
           "RPA30_DataBlock".RPA30_show_points_hmi := 0;
           "RPA30_DataBlock".RPA30_UseInterval_Primer207 := false;
           "RPA30_DataBlock".RPA30_UseIntervalBottleRemover208 := false;
           "RPA30_DataBlock".RPA30_cyclusState := "RPA30_go_to_home_position";
       END_IF;

       "RPA30_DataBlock".RPA30_actual_instruction_index := 255;

       "RPA30R_Beacon_1_LCDPanelGreen" := false;
       "RPA30R_Beacon_1_LCDPanelOrange" := false;
       "RPA30R_Beacon_1_LCDPanelRed" := false;
       "RPA30R_Beacon_1_LCDPanelSiren" := false;
       "RPA30R_Beacon_2_PrimerBoxGreen" := false;
       "RPA30R_Beacon_2_PrimerBoxOrange" := false;
       "RPA30R_Beacon_2_PrimerBoxRed" := false;
       "RPA30R_Beacon_2_PrimerBoxSiren" := false;

       "RPA30R_PrimerPA30GreenReady" := false;
       "RPA30R_PrimerPA30GreenFelt" := false;
       "RPA30R_PrimerPA30GreenRemover208" := false;
       "RPA30R_PrimerPA30GreenPrimer207" := false;
       "RPA30R_PrimerPA30RedNotReady" := false;
       "RPA30R_PrimerPA30RedChangePad" := false;
       "RPA30R_LedBlueConfirm" := false;
       "RPA30R_light" := false;

       "RPA30_DataBlock".RPA30_scannedFrameBareCode := '';

       //if station not active
       "StartStation"(startButton := "RPA30R_LCDButtonStart",
                      StationStartControlVariable := "RPA30_DataBlock".RPA30_Start,
                      stationLight := "RPA30R_light");

       "startButtonLightControlHandler"(stationActivitycontrolVariable := "RPA30_DataBlock".RPA30_Start,
                                        startButtonLED := "RPA30R_LEDGreenSart");
   END_IF;



   IF "RPA30_DataBlock".RPA30_state_information_send = true THEN
       "RPA30_DataBlock".RPA30_state_information_send := NOT "pa30r_station_monitoring"(station_configuration := "RPA30_DataBlock".RPA30_station_configuration,
                                                                                       fail_state := "RPA30_DataBlock".RPA30_failStateLock,
                                                                                       big_fail_state := "RPA30_DataBlock".RPA30_bigFailStateLock,
                                                                                       error_state := "RPA30_DataBlock".RPA30_ErrorStateLock,
                                                                                       fatal_error_state := "RPA30_DataBlock".RPA30_fatalErrorStateLock,
                                                                                       work_cyclus_state := "RPA30_DataBlock".RPA30_actual_instruction_index,
                                                                                       current_frame_code := "RPA30_DataBlock".RPA30_scannedFrameBareCode,
                                                                                       station_activity_state := "RPA30_DataBlock".RPA30_Start,
                                                                                       position_sensor_y := "RPA30R_RoofRotationSensorYAtOperator",
                                                                                       server_connection := "tcp_datablock".tcp_connection,
                                                                                       index:="tcp_datablock".pa30r_station_state_index);
   ELSE
       IF "RPA30_DataBlock".RPA30_fail_state_pre <> "RPA30_DataBlock".RPA30_failStateLock OR
           "RPA30_DataBlock".RPA30_error_state_pre <> "RPA30_DataBlock".RPA30_ErrorStateLock OR
           "RPA30_DataBlock".RPA30_big_fail_state_pre <> "RPA30_DataBlock".RPA30_bigFailStateLock OR
           "RPA30_DataBlock".RPA30_fatal_error_state_pre <> "RPA30_DataBlock".RPA30_fatalErrorStateLock OR
           "RPA30_DataBlock".RPA30_current_frame_code_pre <> "RPA30_DataBlock".RPA30_scannedFrameBareCode OR
           "RPA30_DataBlock".RPA30_hmi_state_pre <> "RPA30_DataBlock".RPA30_actual_instruction_index OR
           "RPA30_DataBlock".RPA30_position_y_pre <> "RPA30R_RoofRotationSensorYAtOperator" OR
           "RPA30_DataBlock".RPA30_station_activity_state_pre <> "RPA30_DataBlock".RPA30_Start THEN

           "RPA30_DataBlock".RPA30_state_information_send := true;
       END_IF;

       "RPA30_DataBlock".RPA30_fail_state_pre := "RPA30_DataBlock".RPA30_failStateLock;
       "RPA30_DataBlock".RPA30_error_state_pre := "RPA30_DataBlock".RPA30_ErrorStateLock;
       "RPA30_DataBlock".RPA30_big_fail_state_pre := "RPA30_DataBlock".RPA30_bigFailStateLock;
       "RPA30_DataBlock".RPA30_fatal_error_state_pre := "RPA30_DataBlock".RPA30_fatalErrorStateLock;
       "RPA30_DataBlock".RPA30_current_frame_code_pre := "RPA30_DataBlock".RPA30_scannedFrameBareCode;
       "RPA30_DataBlock".RPA30_hmi_state_pre := "RPA30_DataBlock".RPA30_actual_instruction_index;
       "RPA30_DataBlock".RPA30_position_y_pre := "RPA30R_RoofRotationSensorYAtOperator";
       "RPA30_DataBlock".RPA30_station_activity_state_pre := "RPA30_DataBlock".RPA30_Start;
   END_IF;
END_FUNCTION

FUNCTION "RPA60_Main" : Void   // FC21, SCL
{ S7_Optimized_Access := 'FALSE' }
VERSION : 0.1
BEGIN
   //main function of station
   IF "RPA60_DataBlock".RPA60_Start = true THEN
       //cyclus handler function
       IF NOT "RPA60R_LCDSwitchAutomat_Manual" THEN

           "server_connection_handler"(error_state_lock_identifier := 1000,
                                       fatal_error_state_lock := "RPA60_DataBlock".RPA60_fatalErrorStateLock,
                                       database_connection := "tcp_datablock".tcp_connection,
                                       error_state_lock := "RPA60_DataBlock".RPA60_ErrorStateLock);

           "RPA60_RollerPresenceHandler"(errorStateLock := "RPA60_DataBlock".RPA60_ErrorStateLock,
                                         fatalErrorStateLock := "RPA60_DataBlock".RPA60_fatalErrorStateLock,
                                         rollerPresenceSensor := "RPA60R_SenzorRoller",
                                         roller_in_use := "RPA60_DataBlock".RPA60_rollerUsageInterval,
                                         roller_taking := "RPA60_DataBlock".RPA60_roller_taking,
                                         bigFailStateIdentifire := 20,
                                         confirmButton := "RPA60R_LCDButtonConfirmSignal",
                                         rollerLED => "RPA60R_LEDRoller",
                                         confirmButtonLed => "RPA60R_LedBlueConfirm",
                                         bigFailStateLock := "RPA60_DataBlock".RPA60_bigFailStateLock,
                                         workCyclusControlVariable := "RPA60_DataBlock".RPA60_cyclusState);
           //*)    

           "RPA60_Scanner_DB"("PORT" := "pa60~CM_PtP_1",
                              BUFFER := "RPA60_Scanner_DB".ReceiveBuffer,
                              NDR => "RPA60_Scanner_DB".NDR,
                              ERROR => "RPA60_Scanner_DB".ERROR,
                              STATUS => "RPA60_Scanner_DB".STATUS,
                              LENGTH => "RPA60_Scanner_DB".LENGTH);

           IF "RPA60_Scanner_DB".NDR = true THEN
               Chars_TO_Strg(Chars := "RPA60_Scanner_DB".ReceiveBuffer,
                             pChars := 0,
                             Cnt := "RPA60_Scanner_DB".received_length - 1,
                             Strg => "RPA60_DataBlock".RPA60_scanedData);
           END_IF;

           "RPA60_HandlerFunction"();




           //beacon light control
           "beaconStateControl"(big_fail_state_lock:="RPA60_DataBlock".RPA60_bigFailStateLock,
                                fail_state_lock:="RPA60_DataBlock".RPA60_failStateLock,
                                error_state_lock:="RPA60_DataBlock".RPA60_ErrorStateLock,
                                fatal_error_state_lock:="RPA60_DataBlock".RPA60_fatalErrorStateLock,
                                beaconGreen := "RPA60R_Beacon_1_LCDPanelGreen",
                                beaconOrange := "RPA60R_Beacon_1_LCDPanelOrange",
                                beaconRed := "RPA60R_Beacon_1_LCDPanelRed");

           //siren control
           "sirenPulsingHandler"(fatal_error:="RPA60_DataBlock".RPA60_fatalErrorStateLock,
                                 big_fail:="RPA60_DataBlock".RPA60_bigFailStateLock,
                                 siren_handler_enable:="RPA60_DataBlock".RPA60_siren_hadler_enable,
                                 siren := "RPA60R_Beacon_1_LCDPanelSiren");




           //valve error checking        
            "valveErrorHandler"(valveLock := "RPA60R_ValveCylinderYLock",
                                valveLockState := "RPA60R_ValveCylinderYLock",
                                valveErrorCheckingState := "RPA60_DataBlock".RPA60_valveYErrorStateCheck,
                                fatalErrorSectionLock := 150,
                                confirmButton := "RPA60R_LCDButtonConfirmSignal",
                                fatalErrorLock := "RPA60_DataBlock".RPA60_fatalErrorStateLock,
                                confirmButtonLED := "RPA60R_LedBlueConfirm");


           //vacuum control
           //
            IF ("RPA60_DataBlock".RPA60_failStateLock + "RPA60_DataBlock".RPA60_bigFailStateLock + "RPA60_DataBlock".RPA60_ErrorStateLock + "RPA60_DataBlock".RPA60_fatalErrorStateLock) = 0 THEN
                "pa60r_vacuum_cleaner_controll_DB"(vacuum_sensor := "RPA60R_SenzorVacuum",
                                                   vacuum_control_variable := "RPA60R_VacuumSwitch");
            END_IF;
       END_IF;
   ELSE
       //if station not active
       IF "lockAxis"(valvePositionSensor := "RPA60R_ValveCylinderYLock",
                         valveNewState := false,
                         valve_error_checking := "RPA60_DataBlock".RPA60_valveYErrorStateCheck,
                         valve := "RPA60R_ValveCylinderYLock") THEN

           "RPA60_DataBlock".RPA60_show_check_button := false;
           "RPA60_DataBlock".RPA60_number_of_check := 0;
           "RPA60_DataBlock".RPA60_bigFailStateLock := 0;
           "RPA60_DataBlock".RPA60_ErrorStateLock := 0;
           "RPA60_DataBlock".RPA60_failStateLock := 0;
           "RPA60_DataBlock".RPA60_fatalErrorStateLock := 0;

           "RPA60_DataBlock".RPA60_printEnable := true;
           "RPA60_DataBlock".RPA60_show_smile := false;
           "RPA60_DataBlock".RPA60_roller_taking := false;
           "RPA60_DataBlock".RPA60_rollerUsageInterval := false;
           "RPA60_DataBlock".RPA60_cyclusState := "RPA60_go_to_home_position";
           "RPA60_DataBlock".RPA60_hmi_instruction_index := 255;
       END_IF;

       "RPA60R_LedBlueConfirm" := false;
       "RPA60R_LEDRoller" := false;
       "RPA60R_Beacon_1_LCDPanelGreen" := false;
       "RPA60R_Beacon_1_LCDPanelOrange" := false;
       "RPA60R_Beacon_1_LCDPanelRed" := false;
       "RPA60R_Beacon_1_LCDPanelSiren" := false;

       "RPA60R_light" := false;

       "StartStation"(startButton := "RPA60R_LCDButtonStart",
                      StationStartControlVariable := "RPA60_DataBlock".RPA60_Start,
                      stationLight := "RPA60R_light");

       "startButtonLightControlHandler"(stationActivitycontrolVariable := "RPA60_DataBlock".RPA60_Start,
                                        startButtonLED := "RPA60R_LEDGreenSart");

   END_IF;

   IF "RPA60_DataBlock".RPA60_state_information_send = true THEN
       "RPA60_DataBlock".RPA60_state_information_send := NOT "pa60r_station_monitoring"(station_configuration:="RPA60_DataBlock".RPA60_station_configuration,
                             fail_state:="RPA60_DataBlock".RPA60_failStateLock,
                             big_fail_state:="RPA60_DataBlock".RPA60_bigFailStateLock,
                             error_state:="RPA60_DataBlock".RPA60_ErrorStateLock,
                             fatal_error_state:="RPA60_DataBlock".RPA60_fatalErrorStateLock,
                             work_cyclus_state:="RPA60_DataBlock".RPA60_hmi_instruction_index,
                             current_frame_code:="RPA60_DataBlock".RPA60_scannedFrameBareCode,
                             station_activity_state:="RPA60_DataBlock".RPA60_Start,
                             position_sensor_y:="RPA60R_RoofRotationSensorYAtOperator",
                             server_connection:="tcp_datablock".tcp_connection, index:="tcp_datablock".pa60r_station_state_index);

   ELSE
       IF "RPA60_DataBlock".RPA60_fail_state_pre <> "RPA60_DataBlock".RPA60_failStateLock OR
           "RPA60_DataBlock".RPA60_error_state_pre <> "RPA60_DataBlock".RPA60_ErrorStateLock OR
           "RPA60_DataBlock".RPA60_big_fail_state_pre <> "RPA60_DataBlock".RPA60_bigFailStateLock OR
           "RPA60_DataBlock".RPA60_fatal_error_state_pre <> "RPA60_DataBlock".RPA60_fatalErrorStateLock OR
           "RPA60_DataBlock".RPA60_current_frame_code_pre <> "RPA60_DataBlock".RPA60_scannedFrameBareCode OR
           "RPA60_DataBlock".RPA60_hmi_state_pre <> "RPA60_DataBlock".RPA60_hmi_instruction_index OR
           "RPA60_DataBlock".RPA60_position_y_pre <> "RPA60R_RoofRotationSensorYAtOperator" OR
           "RPA60_DataBlock".RPA60_station_activity_state_pre <> "RPA60_DataBlock".RPA60_Start THEN
           "RPA60_DataBlock".RPA60_state_information_send := true;
       END_IF;

       "RPA60_DataBlock".RPA60_fail_state_pre := "RPA60_DataBlock".RPA60_failStateLock;
       "RPA60_DataBlock".RPA60_error_state_pre := "RPA60_DataBlock".RPA60_ErrorStateLock;
       "RPA60_DataBlock".RPA60_big_fail_state_pre := "RPA60_DataBlock".RPA60_bigFailStateLock;
       "RPA60_DataBlock".RPA60_fatal_error_state_pre := "RPA60_DataBlock".RPA60_fatalErrorStateLock;
       "RPA60_DataBlock".RPA60_current_frame_code_pre := "RPA60_DataBlock".RPA60_scannedFrameBareCode;
       "RPA60_DataBlock".RPA60_hmi_state_pre := "RPA60_DataBlock".RPA60_hmi_instruction_index;
       "RPA60_DataBlock".RPA60_position_y_pre := "RPA60R_RoofRotationSensorYAtOperator";
       "RPA60_DataBlock".RPA60_station_activity_state_pre := "RPA60_DataBlock".RPA60_Start;
   END_IF;
END_FUNCTION

FUNCTION "setFatalErrorState" : Void   // FC22, SCL
{ S7_Optimized_Access := 'FALSE' }
VERSION : 0.1
BEGIN

   IF #fatalErrorStateLock = 0 OR #fatalErrorStateLock = #identifier THEN
       #fatalErrorStateLock := #identifier;
       #setFatalErrorState := true;
   ELSE
       #setFatalErrorState := false;
   END_IF;
END_FUNCTION

FUNCTION "bottleLightControl" : Void   // FC23, SCL
{ S7_Optimized_Access := 'FALSE' }
VERSION : 0.1
BEGIN

   IF (#failStateLock = 0 OR #failStateLock = #sectionFailIdentifier OR #failStateLock = (#sectionFailIdentifier + 100)) AND
       #bigFailStateLock = 0 AND #ErrorStateLock = 0 AND #FatalErrorStateLock = 0 THEN

       #bottleLight := #bottlePresenceSensor AND "Clock_0.5Hz" AND #bottleInUsage OR (NOT #bottlePresenceSensor);

       IF #failStateLock = #sectionFailIdentifier THEN
           "setOKState"(confirm := true,
                        identifier := #sectionFailIdentifier,
                        confirm_blinking := false,
                        blinkConfirmButton => #buttonConfirmLED,
                        stateLock := #failStateLock);
       ELSE
           "setOKState"(confirm := true,
                        identifier := #sectionFailIdentifier + 100,
                        confirm_blinking := false,
                        blinkConfirmButton => #buttonConfirmLED,
                        stateLock := #failStateLock);
       END_IF;

       IF #bottleInUsage THEN
           IF #bottlePresenceSensor THEN
               IF #bottle_taking THEN
                   IF "setFailState"(identifier := #sectionFailIdentifier, failStateLock := #failStateLock) = true THEN
                       ;
                   END_IF;
               END_IF;
           END_IF;
       ELSE
           IF NOT #bottlePresenceSensor THEN
               IF "setFailState"(identifier := #sectionFailIdentifier+100, failStateLock := #failStateLock) = true THEN
                   ;
               END_IF;
           END_IF;
       END_IF;
   END_IF;
END_FUNCTION

FUNCTION "add_table_record" : Void   // FC25, SCL
{ S7_Optimized_Access := 'FALSE' }
VERSION : 0.1
BEGIN
   #add_table_record := false;

   IF #server_connection = true THEN

       IF #index = 255 THEN
           #msg_out := CONCAT(IN1 := 'SQL~INSERT INTO ', IN2 := #table);
           #msg_out := CONCAT(IN1 := #msg_out, IN2 := ' (');
           Strg_TO_Chars(Strg := #msg_out,
                         pChars := 0,
                         Cnt => #chars,
                         Chars := #temp_buffer);
           #i := #chars;
           #chars := #i;

           WHILE #new_record_items[#i - #chars] <> '$L' AND #i < 1023 DO
               #temp_buffer[#i] := #new_record_items[#i - #chars];
               #i := #i + 1;
           END_WHILE;

           Strg_TO_Chars(Strg := ') VALUES (',
                         pChars := #i,
                         Cnt => #chars,
                         Chars := #temp_buffer);

           #i := #i + #chars;
           #chars := #i;

           WHILE #new_record_data[#i - #chars] <> '$L' AND #i < 1023 DO
               #temp_buffer[#i] := #new_record_data[#i - #chars];
               #i := #i + 1;
           END_WHILE;

           Strg_TO_Chars(Strg := ');$L',
                         pChars := #i,
                         Cnt => #chars,
                         Chars := #temp_buffer);
           #i := #i + #chars;




           #msg_index := "tcp_send"(#temp_buffer);
           IF #msg_index <> 255 THEN
               #index := #msg_index;

           END_IF;
       ELSE
           IF "tcp_rcv"(msg_index := #index, rcv_data => #temp_buffer) = true THEN
               #add_table_record := true;
               #index := 255;
           END_IF;
       END_IF;
   END_IF;
END_FUNCTION

FUNCTION "get_table_record" : Void   // FC26, SCL
{ S7_Optimized_Access := 'FALSE' }
VERSION : 0.1
BEGIN
   #get_table_record := false;

   IF #server_connection = true THEN
       IF #index = 255 THEN
           #msg_out := CONCAT(IN1 := 'GET_TABLE_RECORD', IN2 := '~');
           #msg_out := CONCAT(IN1 := #msg_out, IN2 := #table);
           #msg_out := CONCAT(IN1 := #msg_out, IN2 := '~');
           #msg_out := CONCAT(IN1 := #msg_out, IN2 := #record_key);
           #msg_out := CONCAT(IN1 := #msg_out, IN2 := '~');
           #msg_out := CONCAT(IN1 := #msg_out, IN2 := #record);
           #msg_out := CONCAT(IN1 := #msg_out, IN2 := '$L');

           Strg_TO_Chars(Strg := #msg_out,
                         pChars := 0,
                         Cnt => #chars,
                         Chars := #temp_buffer);

           #msg_index := "tcp_send"(#temp_buffer);
           IF #msg_index <> 255 THEN
               #index := #msg_index;
           END_IF;
       ELSE
           IF "tcp_rcv"(msg_index := #index, rcv_data => #output_buffer) THEN
               #get_table_record := true;
               #index := 255;
           END_IF;
       END_IF;
   END_IF;
END_FUNCTION

FUNCTION "get_table_record_item" : Void   // FC27, SCL
{ S7_Optimized_Access := 'FALSE' }
VERSION : 0.1
BEGIN
   #get_table_record_item := false;

   IF #server_connection = true THEN
       IF #index = 255 THEN
           #msg_out := CONCAT(IN1 := 'GET_TABLE_RECORD_ITEM', IN2 := '~');
           #msg_out := CONCAT(IN1 := #msg_out, IN2 := #table);
           #msg_out := CONCAT(IN1 := #msg_out, IN2 := '~');
           #msg_out := CONCAT(IN1 := #msg_out, IN2 := #record);
           #msg_out := CONCAT(IN1 := #msg_out, IN2 := '~');
           #msg_out := CONCAT(IN1 := #msg_out, IN2 := #item);
           #msg_out := CONCAT(IN1 := #msg_out, IN2 := '~');
           #msg_out := CONCAT(IN1 := #msg_out, IN2 := #record_key);
           #msg_out := CONCAT(IN1 := #msg_out, IN2 := '$L');

           Strg_TO_Chars(Strg := #msg_out,
                         pChars := 0,
                         Cnt => #chars,
                         Chars := #temp_buffer);
           #msg_index := "tcp_send"(#temp_buffer);

           IF #msg_index <> 255 THEN
               #index := #msg_index;
           END_IF;
       ELSE
           IF "tcp_rcv"(msg_index := #index, rcv_data => #output_buffer) = true THEN
               #get_table_record_item := true;
               #index := 255;
           END_IF;
       END_IF;
   END_IF;
END_FUNCTION

FUNCTION "set_table_record_item" : Void   // FC28, SCL
{ S7_Optimized_Access := 'FALSE' }
VERSION : 0.1
BEGIN
       #set_table_record_item := false;

   IF #server_connection = true THEN
       IF #index = 255 THEN
           #msg_out := CONCAT(IN1 := 'SET_TABLE_RECORD_ITEM', IN2 := '~');
           #msg_out := CONCAT(IN1 := #msg_out, IN2 := #table);
           #msg_out := CONCAT(IN1 := #msg_out, IN2 := '~');
           #msg_out := CONCAT(IN1 := #msg_out, IN2 := #record);
           #msg_out := CONCAT(IN1 := #msg_out, IN2 := '~');
           #msg_out := CONCAT(IN1 := #msg_out, IN2 := #record_key);
           #msg_out := CONCAT(IN1 := #msg_out, IN2 := '~');
           #msg_out := CONCAT(IN1 := #msg_out, IN2 := #item);
           #msg_out := CONCAT(IN1 := #msg_out, IN2 := '~');
           #msg_out := CONCAT(IN1 := #msg_out, IN2 := #new_item_data);
           #msg_out := CONCAT(IN1 := #msg_out, IN2 := '$L');

           Strg_TO_Chars(Strg := #msg_out,
                         pChars := 0,
                         Cnt => #chars,
                         Chars := #temp_buffer);

           #msg_index := "tcp_send"(#temp_buffer);

           IF #msg_index <> 255 THEN
               #index := #msg_index;
           END_IF;
       ELSE
           IF "tcp_rcv"(msg_index := #index, rcv_data => #temp_buffer) = true THEN
               #set_table_record_item := true;
               #index := 255;
           END_IF;
       END_IF;
   END_IF;
END_FUNCTION

FUNCTION "startButtonLightControlHandler" : Void   // FC29, SCL
{ S7_Optimized_Access := 'FALSE' }
VERSION : 0.1
BEGIN
   IF #stationActivitycontrolVariable = true THEN
       #startButtonLED := false;
   ELSE
       #startButtonLED := "Clock_0.5Hz";
   END_IF;
END_FUNCTION

FUNCTION "valveErrorHandler" : Void   // FC30, SCL
{ S7_Optimized_Access := 'FALSE' }
VERSION : 0.1
BEGIN

   IF "checkFatalErrorStateLock"(FatalErrorStateLock :=#fatalErrorLock , FatalErrorStatelockIdetifier := #fatalErrorSectionLock) = true
       AND #valveErrorCheckingState = 0 THEN

       IF #valveLock = #valveLockState THEN
           IF #fatalErrorLock = #fatalErrorSectionLock THEN
               "setOKState"(confirm := #confirmButton,
                            identifier := #fatalErrorSectionLock,
                            confirm_blinking := true,
                            blinkConfirmButton => #confirmButtonLED,
                            stateLock := #fatalErrorLock);
           END_IF;
       ELSE
           IF "setFatalErrorState"(identifier := #fatalErrorSectionLock,
                                       fatalErrorStateLock := #fatalErrorLock) THEN
               ;
          END_IF;
       END_IF;

   END_IF;
END_FUNCTION

FUNCTION "lockAxis" : Void   // FC31, SCL
{ S7_Optimized_Access := 'FALSE' }
VERSION : 0.1
BEGIN
   (*
   nastavení pístu do nové polohy, pokud dojde k potvrzení polohy pístu, je vrácena hodnota true
   *)

   #valve := #valveNewState;
   #valve_error_checking := 2000;
   IF #valvePositionSensor = #valveNewState THEN
       #lockAxis := true;
   ELSE
       #lockAxis := false;
   END_IF;
END_FUNCTION

FUNCTION "RPA60_RollerPresenceHandler" : Void   // FC32, SCL
{ S7_Optimized_Access := 'FALSE' }
VERSION : 0.1
BEGIN

   (*
   pokud je big fail state odemčený pak se podprogram vykoná

   pokud přítlačné kolečko ve stavu využíváno pak je rozlišováno jestli se jedná o stav ve kterém se čeká na vyjmutí z dokovací stanice a nebo jestli již je vyjmuto z dokovací stanice

   pokud se jedná o stav kdy se čeká na vyjmutí z dokovací stanice musí blikat světelná kontrolka přítlačného kolečka a být nastaven vnitřní stav stanice OK

   pokud se jedná o stav kdy již je přítlačné kolečko z dokovací stanice vyjmuto kontroluje se zda není vloženo zpátky před expirací časovače

   pokud je přítlačné kolečko vloženo do dokovací stanice před expirací časovače dojde k nastavení stavu big fail a blikání světelné kontrolky přítlačného kolečka

   *)

   IF (#bigFailStateLock = 0 OR #bigFailStateLock = #bigFailStateIdentifire OR #bigFailStateLock = #bigFailStateIdentifire + 100) AND
       #errorStateLock = 0 AND
       #fatalErrorStateLock = 0 THEN

       //blikání a svícení světelné kontrolky přítlačného kolečka
       //#bottlePresenceSensor AND "Clock_0.5Hz" AND #bottleInUsage
       #rollerLED := (NOT #rollerPresenceSensor) OR (#rollerPresenceSensor AND "Clock_0.5Hz" AND #roller_in_use);
       //#rollerLED := (NOT #rollerPresenceSensor) OR (#rollerPresenceSensor AND #rollerUsageInterval[#workCyclusControlVariable] AND "Clock_0.5Hz");

       IF #bigFailStateLock = #bigFailStateIdentifire  THEN
           "setOKState"(confirm := true,
                        identifier := #bigFailStateIdentifire,
                        confirm_blinking := false,
                        blinkConfirmButton => #confirmButtonLed,
                        stateLock := #bigFailStateLock);
       ELSIF #bigFailStateLock = #bigFailStateIdentifire+100 AND #rollerPresenceSensor = true THEN
               "setOKState"(confirm := #confirmButton,
                            identifier := #bigFailStateIdentifire+100,
                            confirm_blinking := true,
                            blinkConfirmButton => #confirmButtonLed,
                            stateLock := #bigFailStateLock);
       END_IF;
       //kontrola přítomnosti kolečka v pracovním cyklu
       IF #roller_in_use THEN
           //nekontroluje první stav a poslední stav ve kterém je přítlačné kolečko používáno -> stav ve kterém se mění mění přítomnost kolečka v dokovací stanici
           IF #roller_in_use THEN
               IF #rollerPresenceSensor THEN
                   IF #roller_taking THEN
                       IF "setBigFailState"(identifier := #bigFailStateIdentifire,
                                                error_state_lock:="RPA60_DataBlock".RPA60_ErrorStateLock, fatal_state_error:="RPA60_DataBlock".RPA60_fatalErrorStateLock, badfailStateLock := #bigFailStateLock) THEN
                           ;
                       END_IF;
                   END_IF;
               END_IF;
           END_IF;
       ELSE
           IF (NOT #rollerPresenceSensor) THEN
               IF "setBigFailState"(identifier := #bigFailStateIdentifire + 100,
                                        error_state_lock:="RPA60_DataBlock".RPA60_ErrorStateLock, fatal_state_error:="RPA60_DataBlock".RPA60_ErrorStateLock, badfailStateLock := #bigFailStateLock) THEN
                   ;
               END_IF;
           END_IF;
       END_IF;
   ELSE
       #rollerLED := false;
   END_IF;
END_FUNCTION

FUNCTION "RPA30_IFM_runtime_switching" : Void   // FC33, SCL
{ S7_Optimized_Access := 'FALSE' }
VERSION : 0.1
BEGIN


   "PA30_IFM_Left_PulsApplicationSwitch_DB"(IFM_Pulse_Period := 15,
                                            IFM_Input_1 := "RPA30R_SensorIFMLeft_Input_1",
                                            IFM_Input_2 := "RPA30R_SensorIFMLeft_Input_2",
                                            ready_intput := "RPA30R_SensorIFMLeftReadyOut");

   "PA30_IFM_Right_PulsApplicationSwitch_DB"(IFM_Pulse_Period := 15,
                                             IFM_Input_1 := "RPA30R_SensorIFMRight_Input_1",
                                             IFM_Input_2 := "RPA30R_SensorIFMRight_Input_2",
                                             ready_intput := "RPA30R_SensorIFMRightReadyOut");
END_FUNCTION

FUNCTION "RPA60_CheckHardwareConfiguration" : Void   // FC34, SCL
{ S7_Optimized_Access := 'FALSE' }
VERSION : 0.1
BEGIN

   CASE #hardwareConfiguration OF
       0:
           #RPA60_CheckHardwareConfiguration := (#senzor_1) AND (NOT #senzor_2);
       1:  
           #RPA60_CheckHardwareConfiguration := (NOT #senzor_1) AND (#senzor_2);
       2:
           #RPA60_CheckHardwareConfiguration := (#senzor_1) AND (#senzor_2);
       ELSE  
           #RPA60_CheckHardwareConfiguration := false;
   END_CASE;
END_FUNCTION

FUNCTION "ping" : Void   // FC35, SCL
{ S7_Optimized_Access := 'FALSE' }
VERSION : 0.1
BEGIN
   #ping := false;

   IF #server_connection = true THEN
       IF "tcp_datablock".ping_index = 255 THEN
           Strg_TO_Chars(Strg := 'PING$L',
                         pChars := 0,
                         Cnt => #chars,
                         Chars := #temp_buffer);

           #index := "tcp_send"(#temp_buffer);

           IF #index <> 255 THEN
               "tcp_datablock".ping_index := #index;
           END_IF;
       ELSE
           IF "tcp_rcv"(msg_index := "tcp_datablock".ping_index, rcv_data => #temp_buffer) = true THEN
               IF "parse_input_data"(#temp_buffer) = 'OK' THEN
                   #server_connection := true;
               ELSE
                   #server_connection := false;
               END_IF;
               #ping := true;
               "tcp_datablock".ping_index := 255;
           END_IF;
       END_IF;
   END_IF;
END_FUNCTION

FUNCTION "setFailState" : Void   // FC36, SCL
{ S7_Optimized_Access := 'FALSE' }
VERSION : 0.1
BEGIN

   IF #failStateLock = 0 OR #failStateLock = #identifier THEN
       #failStateLock := #identifier;
       #setFailState := true;
   ELSE
       #setFailState := false;
   END_IF;
END_FUNCTION

FUNCTION "bottle_label_check" : Void   // FC37, SCL
{ S7_Optimized_Access := 'FALSE' }
VERSION : 0.1
BEGIN
   (*
    * formát dat: kód chemikálie*batch kód*filling date*expire date*druh lahvičky*identifikátor stanice
    * každá část je oddělena znakem '*'
    *)

   #bottle_label_check := 0;
   IF #chemical_type > 0 AND #chemical_type < 6 THEN
       (* parse input date *)
       #index := 1;
       #part := 0;
       WHILE #index <= LEN(#input_data) DO
           IF #input_data[#index] = '*' THEN
               #part := #part + 1;
           ELSE
               CASE #part OF
                   0: 
                       #chemical_code := CONCAT(IN1 := #chemical_code, IN2 := #input_data[#index]);
                   2:
                       #expiring_date_time := CONCAT(IN1 := #expiring_date_time, IN2 := #input_data[#index]);
                   5:
                       #bottle_type := CONCAT(IN1 := #bottle_type, IN2 := #input_data[#index]);
               END_CASE;
           END_IF;

           #index := #index +1;
       END_WHILE;

           (* check chemical *)
           IF (#chemical_type = 1 AND #chemical_code = '1714290C') OR
               (#chemical_type = 2 AND #chemical_code = '1714291A') OR
               (#chemical_type = 3 AND #chemical_code = '1704681') OR
               (#chemical_type = 4 AND #chemical_code = '1742250B') OR
               (#chemical_type = 5 AND #chemical_code = '17422749') THEN

               (* checking bottle type *)
               IF #bottle_type = 'S' THEN
                   (* check expiration date *)
                   #expire_date_time.DAY := STRING_TO_USINT("sub_string"(str_in := #expiring_date_time, start_index := 1, end_index := 2));
                   #expire_date_time.MONTH := STRING_TO_USINT("sub_string"(str_in := #expiring_date_time, start_index := 4, end_index := 5));
                   #expire_date_time.YEAR := STRING_TO_UINT("sub_string"(str_in := #expiring_date_time, start_index := 7, end_index := 10));

                   #expire_date_time.HOUR := STRING_TO_USINT("sub_string"(str_in := #expiring_date_time, start_index := 12, end_index := 13));
                   #expire_date_time.MINUTE := STRING_TO_USINT("sub_string"(str_in := #expiring_date_time, start_index := 15, end_index := 16));

                   IF RD_SYS_T(#current_date_time) < 2 THEN
                       ;
                   END_IF;

                   IF "time_compare"(time_1:=#expire_date_time, time_2:=#current_date_time, difference_treshold:=LT#0s) = true THEN
                       #bottle_label_check := 0;
                   ELSE
                       #bottle_label_check := 5;
                   END_IF;
               ELSE
                   #bottle_label_check := 3;
               END_IF;

           ELSE
               #bottle_label_check := 2;
           END_IF;
       ELSE
           #bottle_label_check := 4;
       END_IF;
END_FUNCTION

FUNCTION "remove_record" : Void   // FC38, SCL
{ S7_Optimized_Access := 'FALSE' }
VERSION : 0.1
BEGIN
   #remove_record := false;

   IF #server_connection = true THEN
       IF #index = 255 THEN
           #msg_out := CONCAT(IN1 := 'REMOVE_TABLE_RECORD', IN2 := '~');
           #msg_out := CONCAT(IN1 := #msg_out, IN2 := #table);
           #msg_out := CONCAT(IN1 := #msg_out, IN2 := '~');
           #msg_out := CONCAT(IN1 := #msg_out, IN2 := #record_key);
           #msg_out := CONCAT(IN1 := #msg_out, IN2 := '~');
           #msg_out := CONCAT(IN1 := #msg_out, IN2 := #record);
           #msg_out := CONCAT(IN1 := #msg_out, IN2 := '$L');
           Strg_TO_Chars(Strg := #msg_out,
                         pChars := 0,
                         Cnt => #chars,
                         Chars := #temp_buffer);

           #msg_index := "tcp_send"(#temp_buffer);

           IF #msg_index <> 255 THEN
               #index := #msg_index;
           END_IF;
       ELSE
           IF "tcp_rcv"(msg_index := #index, rcv_data => #temp_buffer) = true THEN
               #remove_record := true;
               #index := 255;
           END_IF;
       END_IF;
   END_IF;
END_FUNCTION

FUNCTION "setBigFailState" : Void   // FC39, SCL
{ S7_Optimized_Access := 'FALSE' }
VERSION : 0.1
BEGIN

   IF #badfailStateLock = 0 OR #badfailStateLock = #identifier AND (#error_state_lock + #fatal_state_error) = 0 THEN
       #badfailStateLock := #identifier;
       #setBigFailState := true;
   ELSE
       #setBigFailState := false;
   END_IF;
END_FUNCTION

FUNCTION "feltLightControl" : Void   // FC40, SCL
{ S7_Optimized_Access := 'FALSE' }
VERSION : 0.1
BEGIN

   IF "checkFailStateLock"(failStateLock:=#failStateLock,
                               bigFailStateLock:=#bigFailStateLock,
                               ErrorStateLock:=#ErrorStateLock,
                               FatalErrorStateLock:=#FatalErrorStateLock,
                               failStatelockIdetifier:=#failStateLockIdentifier) THEN

       IF #feltPresenceSensor = false THEN
           IF "setFailState"(identifier := #failStateLockIdentifier,
                                 failStateLock := #failStateLock) THEN
               ;
           END_IF;
       END_IF;

       #feltLED := NOT #feltPresenceSensor;
       #readyLED := #feltPresenceSensor;
       #notReady := #feltLED;

       IF #failStateLockIdentifier = #failStateLock AND #feltPresenceSensor THEN
           "setOKState"(confirm:=true,
                        identifier:=#failStateLockIdentifier,
                        confirm_blinking:=false,
                        blinkConfirmButton=>#confirmButtonLED,
                        stateLock:=#failStateLock);
       END_IF;
   END_IF;
END_FUNCTION

FUNCTION "setErrorState" : Void   // FC41, SCL
{ S7_Optimized_Access := 'FALSE' }
VERSION : 0.1
BEGIN
   IF #ErrorStateLock = 0 OR #ErrorStateLock = #identifier THEN

       #ErrorStateLock := #identifier;
       #setErrorState := true;
   ELSE
       #setErrorState := false;
   END_IF;
END_FUNCTION

FUNCTION "pa30r_station_monitoring" : Void   // FC42, SCL
{ S7_Optimized_Access := 'FALSE' }
VERSION : 0.1
BEGIN
   #pa30r_station_monitoring := false;
   IF #server_connection = true THEN
       IF #index = 255 THEN
       (* command *)
           Strg_TO_Chars(Strg := 'PA30R_STATE~',
                         pChars := 0,
                         Cnt => #chars,
                         Chars := #temp_buffer);
           #i := #chars;

           (* station state *)
           IF #station_activity_state = true THEN
               IF #fatal_error_state > 0 THEN
                   CASE #fatal_error_state OF
                       150:
                           Strg_TO_Chars(Strg := '<html>Station state: Y axis<br>valve lock error</html>~',
                                         pChars := #i,
                                         Cnt => #chars,
                                         Chars := #temp_buffer);
                       160:
                           Strg_TO_Chars(Strg := 'Station state: Bad frame code~',
                                         pChars := #i,
                                         Cnt => #chars,
                                         Chars := #temp_buffer);
                       ELSE
                           Strg_TO_Chars(Strg := 'Station state: Unknown~',
                                         pChars := #i,
                                         Cnt => #chars,
                                         Chars := #temp_buffer);
                   END_CASE;
               ELSE
                   IF #error_state > 0 THEN
                       CASE #error_state OF
                           22000:
                               Strg_TO_Chars(Strg := 'Station state: Frame already processed~',
                                             pChars := #i,
                                             Cnt => #chars,
                                             Chars := #temp_buffer);
                           23000:
                               Strg_TO_Chars(Strg := 'Station state: More then 8 hours~',
                                             pChars := #i,
                                             Cnt => #chars,
                                             Chars := #temp_buffer);
                           24000:
                               Strg_TO_Chars(Strg := 'Station state: Less then 10 minutes~',
                                             pChars := #i,
                                             Cnt => #chars,
                                             Chars := #temp_buffer);
                           25000:
                               Strg_TO_Chars(Strg := 'Station state: Frame is not in database~',
                                             pChars := #i,
                                             Cnt => #chars,
                                             Chars := #temp_buffer);
                           26000:
                               Strg_TO_Chars(Strg := 'Station state: Bad station configuration~',
                                             pChars := #i,
                                             Cnt => #chars,
                                             Chars := #temp_buffer);
                           ELSE
                               Strg_TO_Chars(Strg := 'Station state: Unknown~',
                                             pChars := #i,
                                             Cnt => #chars,
                                             Chars := #temp_buffer);
                       END_CASE;


                   ELSE
                       IF #big_fail_state > 0 THEN
                           Strg_TO_Chars(Strg := 'Station state: Unknown~',
                                         pChars := #i,
                                         Cnt => #chars,
                                         Chars := #temp_buffer);
                       ELSE
                           IF #fail_state > 0 THEN
                               CASE #fail_state OF
                                   6:
                                       Strg_TO_Chars(Strg := 'Station state: Bottle expiration~',
                                                     pChars := #i,
                                                     Cnt => #chars,
                                                     Chars := #temp_buffer);
                                   300:
                                       Strg_TO_Chars(Strg := 'Station state: Felt box is empty~',
                                                     pChars := #i,
                                                     Cnt => #chars,
                                                     Chars := #temp_buffer);
                                   200:
                                       Strg_TO_Chars(Strg := 'Station state: Primer 207 out of primer box~',
                                                     pChars := #i,
                                                     Cnt => #chars,
                                                     Chars := #temp_buffer);
                                   210:
                                       Strg_TO_Chars(Strg := 'Station state: Remover out of primer box~',
                                                     pChars := #i,
                                                     Cnt => #chars,
                                                     Chars := #temp_buffer);
                                   100:
                                       Strg_TO_Chars(Strg := 'Station state: Primer 207 in primer box~',
                                                     pChars := #i,
                                                     Cnt => #chars,
                                                     Chars := #temp_buffer);
                                   33:
                                       Strg_TO_Chars(Strg := 'Station state: Remover 208 expired~',
                                                     pChars := #i,
                                                     Cnt => #chars,
                                                     Chars := #temp_buffer);
                                   ELSE  // Statement section ELSE
                                       Strg_TO_Chars(Strg := 'Station state: Unknown~',
                                                     pChars := #i,
                                                     Cnt => #chars,
                                                     Chars := #temp_buffer);
                               END_CASE;

                           ELSE
                               Strg_TO_Chars(Strg := 'Station state: OK~',
                                             pChars := #i,
                                             Cnt => #chars,
                                             Chars := #temp_buffer);
                           END_IF;
                       END_IF;
                   END_IF;
               END_IF;
           ELSE
               Strg_TO_Chars(Strg := 'Station state: Inactive~',
                             pChars := #i,
                             Cnt => #chars,
                             Chars := #temp_buffer);
           END_IF;

           #i := #i + #chars;

           (* work cyclus state *)

           IF #work_cyclus_state = "RPA30_hmi_go_to_home_position" THEN
               Strg_TO_Chars(Strg := 'Work cyclus state: Waiting for home position~',
                             pChars := #i,
                             Cnt => #chars,
                             Chars := #temp_buffer);
           ELSIF #work_cyclus_state = "RPA30_hmi_scan_frame" THEN
               Strg_TO_Chars(Strg := 'Work cyclus state: Scan frame code~',
                             pChars := #i,
                             Cnt => #chars,
                             Chars := #temp_buffer);
           ELSIF #work_cyclus_state = "RPA30_hmi_turn_frame_clockwise" THEN
               Strg_TO_Chars(Strg := '<html>Work cyclus state: Turn the frame<br>for 90° clockwise</html>~',
                             pChars := #i,
                             Cnt => #chars,
                             Chars := #temp_buffer);
           ELSIF #work_cyclus_state = "RPA30_hmi_take_felt" THEN
               Strg_TO_Chars(Strg := 'Work cyclus state: Take felt from primer box~',
                             pChars := #i,
                             Cnt => #chars,
                             Chars := #temp_buffer);
           ELSIF #work_cyclus_state = "RPA30_hmi_on_felt_apply_remover" THEN
               Strg_TO_Chars(Strg := 'Work cyclus state: On felt apply remover 208~',
                             pChars := #i,
                             Cnt => #chars,
                             Chars := #temp_buffer);
           ELSIF #work_cyclus_state = "RPA30_hmi_apply_remover_on_5_points" THEN
               Strg_TO_Chars(Strg := 'Work cyclus state: Apply remover 208 on frame~',
                             pChars := #i,
                             Cnt => #chars,
                             Chars := #temp_buffer);
           ELSIF #work_cyclus_state = "RPA30_hmi_turn_frame_counterclockwise" THEN
               Strg_TO_Chars(Strg := 'Work cyclus state: Turn frame counterclockwise~',
                             pChars := #i,
                             Cnt => #chars,
                             Chars := #temp_buffer);
           ELSIF #work_cyclus_state = "RPA30_hmi_apply_primer_on_5_points" THEN
               Strg_TO_Chars(Strg := '<html>Work cyclus state: Apply primer 207<br>on frame</html>~',
                             pChars := #i,
                             Cnt => #chars,
                             Chars := #temp_buffer);
           ELSIF #work_cyclus_state = "RPA30_hmi_scan_primer_bottle" THEN
               Strg_TO_Chars(Strg := 'Work cyclus state: Scan primer 207 bottle~',
                             pChars := #i,
                             Cnt => #chars,
                             Chars := #temp_buffer);
           ELSIF #work_cyclus_state = "RPA30_hmi_take_bottle_of_primer" THEN
               Strg_TO_Chars(Strg := 'Work cyclus state: Take bottle of primer 207 from primer box~',
                             pChars := #i,
                             Cnt => #chars,
                             Chars := #temp_buffer);
           ELSIF #work_cyclus_state = "RPA30_hmi_change_pad" THEN
               Strg_TO_Chars(Strg := 'Work cyclus state: Change pad~',
                             pChars := #i,
                             Cnt => #chars,
                             Chars := #temp_buffer);
           ELSIF #work_cyclus_state = "RPA30_hmi_put_primer_bottle_back" THEN
               Strg_TO_Chars(Strg := '<html>Work cyclus state: Put primer 207 bottle<br>back to primer box</hmtl>~',
                             pChars := #i,
                             Cnt => #chars,
                             Chars := #temp_buffer);
           ELSIF #work_cyclus_state = "RPA30_hmi_end_of_cyclus" THEN
               Strg_TO_Chars(Strg := 'Work cyclus state: End of work cyclus~',
                             pChars := #i,
                             Cnt => #chars,
                             Chars := #temp_buffer);
           ELSIF #work_cyclus_state = "RPA30_hmi_wipe_off" THEN
               Strg_TO_Chars(Strg := 'Work cyclus state: Whipe off~',
                             pChars := #i,
                             Cnt => #chars,
                             Chars := #temp_buffer);
           ELSIF #work_cyclus_state = "RPA30_hmi_scan_remover_bottle" THEN
               Strg_TO_Chars(Strg := 'Work cyclus state: Scan remover 208 bottle~',
                             pChars := #i,
                             Cnt => #chars,
                             Chars := #temp_buffer);
           ELSE
               Strg_TO_Chars(Strg := 'Work cyclus state: Unknown~',
                             pChars := #i,
                             Cnt => #chars,
                             Chars := #temp_buffer);
           END_IF;

           #i := #i + #chars;
           (* home position *)
           IF #position_sensor_y THEN
               Strg_TO_Chars(Strg := 'Home position: Yes~',
                             pChars := #i,
                             Cnt => #chars,
                             Chars := #temp_buffer);
           ELSE
               Strg_TO_Chars(Strg := 'Home position: No~',
                             pChars := #i,
                             Cnt => #chars,
                             Chars := #temp_buffer);
           END_IF;

           #i := #i + #chars;
           (* current frame code *)
           Strg_TO_Chars(Strg := 'Current frame code: ',
                         pChars := #i,
                         Cnt => #chars,
                         Chars := #temp_buffer);
           #i := #i + #chars;
           IF #current_frame_code <> '' THEN
               Strg_TO_Chars(Strg := #current_frame_code,
                             pChars := #i,
                             Cnt => #chars,
                             Chars := #temp_buffer);
           ELSE
               Strg_TO_Chars(Strg := 'None',
                             pChars := #i,
                             Cnt => #chars,
                             Chars := #temp_buffer);
           END_IF;
           #i := #i + #chars;

           (* station configuration *)
           IF #station_configuration = 0 THEN
               Strg_TO_Chars(Strg := '~Station configuration: 581A~',
                             pChars := #i,
                             Cnt => #chars,
                             Chars := #temp_buffer);
           ELSIF #station_configuration = 1 THEN
               Strg_TO_Chars(Strg := '~Station configuration: 581B~',
                             pChars := #i,
                             Cnt => #chars,
                             Chars := #temp_buffer);
           ELSIF #station_configuration = 2 THEN
               Strg_TO_Chars(Strg := '~Station configuration: 582A~',
                             pChars := #i,
                             Cnt => #chars,
                             Chars := #temp_buffer);
           ELSIF #station_configuration = 3 THEN
               Strg_TO_Chars(Strg := '~Station configuration: 582B~',
                             pChars := #i,
                             Cnt => #chars,
                             Chars := #temp_buffer);
           END_IF;

           #i := #i + #chars;
           #temp_buffer[#i] := '$L';
           #msg_index := "tcp_send"(#temp_buffer);
           IF #msg_index <> 255 THEN
               #index := #msg_index;
           END_IF;
       ELSE
           IF "tcp_rcv"(msg_index := #index, rcv_data => #temp_buffer) = true THEN
               #index := 255;
               #pa30r_station_monitoring := true;
           END_IF;
       END_IF;
   END_IF;
END_FUNCTION

